Template "Plantilla-Alta-Sec" 1280x800
   Button "Plantilla_6" at 1196,741 size 81x58; TextOff 'Reconocer'; PictureOff "Asleep Check Mark Icon - Sleep Aid Records_2"
      on Press: SetBit("ReconocerTODAS")
      on Release: ResetBit("ReconocerTODAS")
      Appearance <- "AlarmaNueva"
   GraphicView "Plantilla_Visor de gráficos_17" at 4,4 size 87x38; Picture "logo4"
   Button "Plantilla_7" at 479,748 size 78x50; TextOff 'Compres.'
      on Click: ActivateScreen("MTA-CompBAJA", 0)
   Button "Plantilla_8" at 161,748 size 78x50; TextOff 'Torres'
      on Release: ActivateScreen("MTA-TorresCH", 0)
   Button "Plantilla_9" at 81,748 size 78x50; TextOff 'General'; TextOn 'NavigateHome'; PictureOff "NavigateHome_HMI_1"; PictureOn "NavigateHome_HMI_1"
      on Press: ResetBit("VerCh1MTA"); ResetBit("VerCh2MTA"); ResetBit("VerCh3MTA"); ResetBit("VerCh4MTA")
      on Release: ActivateScreen("MTA-Chillers-General", 0)
   Button "Plantilla_12" at 638,748 size 78x50; TextOff 'Luz'; PictureOff "Lamp2_1"
      on Click: ActivateScreen("IluminaciónMTA", 0)
      Appearance <- "MantenerON"
   Button "Plantilla_13" at 400,748 size 78x50; TextOff 'Torres'
      on Click: ActivateScreen("MTA-TorresCAV", 0)
   Button "Plantilla_14" at 321,748 size 78x50; TextOff 'Secadores'
      on Click: ActivateScreen("MTA-SecALTA", 0)
   Button "Plantilla_15" at 558,748 size 78x50; TextOff 'Secadores'
      on Click: ActivateScreen("MTA-SecBaja", 0)
   Button "Plantilla_16" at 241,748 size 78x50; TextOff 'Compres.'
      on Click: ActivateScreen("MTA-CompALTA", 0)
   Button "Plantilla_17" at 1,740 size 78x58; TextOff 'NavigateHome'; PictureOff "NavigateHome_HMI_1"; PictureOn "NavigateHome_HMI_1"
      on Release: ActivateScreen("INICIO", 0)
   GraphicView "Plantilla_Visor de gráficos_1" at 80,740 size 78x6; Picture "indGris"
   GraphicView "Plantilla_Visor de gráficos_2" at 160,740 size 78x6; Picture "indGris"
   GraphicView "Plantilla_Visor de gráficos_3" at 478,740 size 78x6; Picture "indGris"
   GraphicView "Plantilla_Visor de gráficos_4" at 240,740 size 78x6; Picture "indGris"
   GraphicView "Plantilla_Visor de gráficos_5" at 557,740 size 78x6; Picture "indGris"
   GraphicView "Plantilla_Visor de gráficos_6" at 320,740 size 78x6; Picture "indGris"
   GraphicView "Plantilla_Visor de gráficos_7" at 399,740 size 78x6; Picture "indGris"
   GraphicView "Plantilla_Visor de gráficos_11" at 637,740 size 78x6; Picture "indGris"
   GraphicView "Plantilla_Visor de gráficos_8" at 80,740 size 78x6; Picture "indAmarillo"
      Visibility <- "IndCh"
   GraphicView "Plantilla_Visor de gráficos_9" at 160,740 size 78x6; Picture "indAmarillo"
      Visibility <- "IndTrCh"
   GraphicView "Plantilla_Visor de gráficos_10" at 478,740 size 78x6; Picture "indAmarillo"
      Visibility <- "IndCmpBaja"
   GraphicView "Plantilla_Visor de gráficos_12" at 240,740 size 78x6; Picture "indAmarillo"
      Visibility <- "IndCmpAlta"
   GraphicView "Plantilla_Visor de gráficos_13" at 557,740 size 78x6; Picture "indAmarillo"
      Visibility <- "IndSecBaja"
   GraphicView "Plantilla_Visor de gráficos_14" at 320,740 size 78x6; Picture "indAmarillo"
      Visibility <- "IndSecAlta"
   GraphicView "Plantilla_Visor de gráficos_15" at 399,740 size 78x6; Picture "indAmarillo"
      Visibility <- "IndTrCav"
   GraphicView "Plantilla_Visor de gráficos_16" at 637,740 size 78x6; Picture "indAmarillo"
      Visibility <- "MantenerON"
   TextField "Plantilla_Campo de texto_2" at 521,711 size 69x18; Text 'Baja Presión'
   TextField "Plantilla_Campo de texto_4" at 323,711 size 68x18; Text 'Alta Presión'
   TextField "Plantilla_Campo de texto_3" at 139,711 size 40x18; Text 'Chillers'
   Button "Plantilla_3" at 717,748 size 78x50; TextOff 'Text'; PictureOff "Rayo"
      on Click: ActivateScreen("SentronPAC-MTA", 0)
   Button "Plantilla_5" at 957,748 size 78x50; TextOff 'Text'
   Button "Plantilla_11" at 797,748 size 78x50; TextOff 'Variables Analóg.'
      on Click: ActivateScreen("Grafica", 0)
   GraphicView "Plantilla_Visor de gráficos_18" at 717,740 size 78x6; Picture "indGris"
   GraphicView "Plantilla_Visor de gráficos_19" at 797,740 size 78x6; Picture "indGris"
   GraphicView "Plantilla_Visor de gráficos_20" at 877,740 size 78x6; Picture "indGris"
   GraphicView "Plantilla_Visor de gráficos_21" at 957,740 size 78x6; Picture "indGris"
   GraphicView "Plantilla_Visor de gráficos_22" at 1037,740 size 78x6; Picture "indGris"
   GraphicView "Plantilla_Visor de gráficos_23" at 1037,740 size 78x6; Picture "indAmarillo"
      Visibility <- "AnularSirenaCav"
   Button "Plantilla_1" at 1037,749 size 78x50; TextOff 'Anular Sirena'
      on Click: SetBit("AnularSirena?")
   Button "Plantilla_2" at 1117,741 size 78x58; TextOff 'Avisos'
      on Click: ActivateScreen("MTA-Avisos", 0)
   Button "Plantilla_4" at 877,748 size 78x50; TextOff 'Text'
   GraphicView "Plantilla_Visor de gráficos_24" at 877,740 size 78x6; Picture "indGris"
   GraphicView "Plantilla_Visor de gráficos_25" at 877,740 size 78x6; Picture "indGris"
      Visibility <- "AlarmaBoosters"
   Group "Group" at 1,716 size 1276x84
   GraphicView "Plantilla_Visor de gráficos_26" at 68,9 size 91x26; Picture "eProC logo 4 b"
   GraphicView "Plantilla_Visor de gráficos_27" at 9,8 size 49x29; Picture "eProC logo 4 a"
   GraphicIOField "Campo ES gráfico_4" at 981,258 size 280x222; PictureList "Secador1"
      ProcessValue <- "AnimaMS050"
   GraphicView "Visor de gráficos_4" at 999,137 size 234x314; Picture "secador4"
   GraphicView "Visor de gráficos_15" at 999,137 size 234x314; Picture "secador4d_1"
      Visibility <- "MantMS050"
   GraphicIOField "Campo ES gráfico_8" at 571,212 size 366x99; PictureList "Secador2"
      ProcessValue <- "AnimaMS053"
   GraphicView "Visor de gráficos_3" at 592,100 size 363x184; Picture "secador2_3"
   GraphicView "Visor de gráficos_5" at 592,100 size 363x184; Picture "secador2m_1"
      Visibility <- "MantMS053"
   GraphicIOField "Campo ES gráfico_7" at 674,357 size 309x81; PictureList "Secador2"
      ProcessValue <- "AnimaMS052"
   GraphicView "Visor de gráficos_2" at 696,255 size 292x158; Picture "secador3_1"
   GraphicView "Visor de gráficos_6" at 695,255 size 294x158; Picture "secador3d_1"
      Visibility <- "MantMS052"
   GraphicIOField "Campo ES gráfico_6" at 765,490 size 338x86; PictureList "Secador2"
      ProcessValue <- "AnimaMS051"
   GraphicView "Visor de gráficos_1" at 786,405 size 292x142; Picture "secador3_3"
   GraphicView "Visor de gráficos_14" at 786,405 size 292x142; Picture "secador3d_2"
      Visibility <- "MantMS051"
   Rectangle "Plantilla_Rectángulo_1" at 1,716 size 1276x84
      Visibility <- "AnularSirena?"
   TextField "Plantilla_Campo de texto_5" at 32,732 size 696x50; Text '¿Está seguro de ANULAR la sirena? Si decide anular el sistema dejará de emitir avisos sonoros de manera permanente'
      Visibility <- "AnularSirena?"
   Button "Plantilla_Botón_1" at 1232,724 size 37x34; TextOff 'x'
      on Click: ResetBit("AnularSirena?")
      Visibility <- "AnularSirena?"
   Button "Plantilla_Botón_2" at 945,735 size 112x46; TextOff 'Activar'
      on Click: ResetBit("AnularSirenaCav")
      Visibility <- "AnularSirena?"
      Appearance <- "AnularSirenaCav"
   Button "Plantilla_Botón_3" at 1065,735 size 112x46; TextOff 'Desactivar'
      on Click: SetBit("AnularSirenaCav")
      Visibility <- "AnularSirena?"
      Appearance <- "AnularSirenaCav"
   Switch "Interruptor_1" at 640,315 size 40x40; TextOn '1'; TextOff '0'; CaptionText 'Switch'; PictureOff "MECH2"; PictureOn "MECH1"
      ProcessValue <- "MantMS052"
   Switch "Interruptor_2" at 731,440 size 40x40; TextOn '1'; TextOff '0'; CaptionText 'Switch'; PictureOff "MECH2"; PictureOn "MECH1"
      ProcessValue <- "MantMS051"
   Switch "Interruptor_3" at 540,176 size 40x40; TextOn '1'; TextOff '0'; CaptionText 'Switch'; PictureOff "MECH2"; PictureOn "MECH1"
      ProcessValue <- "MantMS053"
   Switch "Interruptor_4" at 1212,488 size 40x40; TextOn '1'; TextOff '0'; CaptionText 'Switch'; PictureOff "MECH2"; PictureOn "MECH1"
      ProcessValue <- "MantMS050"

Template "Plantilla-Baja-Cmp" 1280x800
   Button "Plantilla_6" at 1196,741 size 81x58; TextOff 'Reconocer'; PictureOff "Asleep Check Mark Icon - Sleep Aid Records_2"
      on Press: SetBit("ReconocerTODAS")
      on Release: ResetBit("ReconocerTODAS")
      Appearance <- "AlarmaNueva"
   GraphicView "Plantilla_Visor de gráficos_17" at 4,4 size 87x38; Picture "logo4"
   Button "Plantilla_7" at 479,748 size 78x50; TextOff 'Compres.'
      on Click: ActivateScreen("MTA-CompBAJA", 0)
   Button "Plantilla_8" at 161,748 size 78x50; TextOff 'Torres'
      on Release: ActivateScreen("MTA-TorresCH", 0)
   Button "Plantilla_9" at 81,748 size 78x50; TextOff 'General'; TextOn 'NavigateHome'; PictureOff "NavigateHome_HMI_1"; PictureOn "NavigateHome_HMI_1"
      on Press: ResetBit("VerCh1MTA"); ResetBit("VerCh2MTA"); ResetBit("VerCh3MTA"); ResetBit("VerCh4MTA")
      on Release: ActivateScreen("MTA-Chillers-General", 0)
   Button "Plantilla_12" at 638,748 size 78x50; TextOff 'Luz'; PictureOff "Lamp2_1"
      on Click: ActivateScreen("IluminaciónMTA", 0)
      Appearance <- "MantenerON"
   Button "Plantilla_13" at 400,748 size 78x50; TextOff 'Torres'
      on Click: ActivateScreen("MTA-TorresCAV", 0)
   Button "Plantilla_14" at 321,748 size 78x50; TextOff 'Secadores'
      on Click: ActivateScreen("MTA-SecALTA", 0)
   Button "Plantilla_15" at 558,748 size 78x50; TextOff 'Secadores'
      on Click: ActivateScreen("MTA-SecBaja", 0)
   Button "Plantilla_16" at 241,748 size 78x50; TextOff 'Compres.'
      on Click: ActivateScreen("MTA-CompALTA", 0)
   Button "Plantilla_17" at 1,740 size 78x58; TextOff 'NavigateHome'; PictureOff "NavigateHome_HMI_1"; PictureOn "NavigateHome_HMI_1"
      on Release: ActivateScreen("INICIO", 0)
   GraphicView "Plantilla_Visor de gráficos_1" at 80,740 size 78x6; Picture "indGris"
   GraphicView "Plantilla_Visor de gráficos_2" at 160,740 size 78x6; Picture "indGris"
   GraphicView "Plantilla_Visor de gráficos_3" at 478,740 size 78x6; Picture "indGris"
   GraphicView "Plantilla_Visor de gráficos_4" at 240,740 size 78x6; Picture "indGris"
   GraphicView "Plantilla_Visor de gráficos_5" at 557,740 size 78x6; Picture "indGris"
   GraphicView "Plantilla_Visor de gráficos_6" at 320,740 size 78x6; Picture "indGris"
   GraphicView "Plantilla_Visor de gráficos_7" at 399,740 size 78x6; Picture "indGris"
   GraphicView "Plantilla_Visor de gráficos_11" at 637,740 size 78x6; Picture "indGris"
   GraphicView "Plantilla_Visor de gráficos_8" at 80,740 size 78x6; Picture "indAmarillo"
      Visibility <- "IndCh"
   GraphicView "Plantilla_Visor de gráficos_9" at 160,740 size 78x6; Picture "indAmarillo"
      Visibility <- "IndTrCh"
   GraphicView "Plantilla_Visor de gráficos_10" at 478,740 size 78x6; Picture "indAmarillo"
      Visibility <- "IndCmpBaja"
   GraphicView "Plantilla_Visor de gráficos_12" at 240,740 size 78x6; Picture "indAmarillo"
      Visibility <- "IndCmpAlta"
   GraphicView "Plantilla_Visor de gráficos_13" at 557,740 size 78x6; Picture "indAmarillo"
      Visibility <- "IndSecBaja"
   GraphicView "Plantilla_Visor de gráficos_14" at 320,740 size 78x6; Picture "indAmarillo"
      Visibility <- "IndSecAlta"
   GraphicView "Plantilla_Visor de gráficos_15" at 399,740 size 78x6; Picture "indAmarillo"
      Visibility <- "IndTrCav"
   GraphicView "Plantilla_Visor de gráficos_16" at 637,740 size 78x6; Picture "indAmarillo"
      Visibility <- "MantenerON"
   TextField "Plantilla_Campo de texto_2" at 521,711 size 69x18; Text 'Baja Presión'
   TextField "Plantilla_Campo de texto_4" at 323,711 size 68x18; Text 'Alta Presión'
   TextField "Plantilla_Campo de texto_3" at 139,711 size 40x18; Text 'Chillers'
   Button "Plantilla_3" at 717,748 size 78x50; TextOff 'Text'; PictureOff "Rayo"
      on Click: ActivateScreen("SentronPAC-MTA", 0)
   Button "Plantilla_5" at 957,748 size 78x50; TextOff 'Text'
   Button "Plantilla_11" at 797,748 size 78x50; TextOff 'Variables Analóg.'
      on Click: ActivateScreen("Grafica", 0)
   GraphicView "Plantilla_Visor de gráficos_18" at 717,740 size 78x6; Picture "indGris"
   GraphicView "Plantilla_Visor de gráficos_19" at 797,740 size 78x6; Picture "indGris"
   GraphicView "Plantilla_Visor de gráficos_20" at 877,740 size 78x6; Picture "indGris"
   GraphicView "Plantilla_Visor de gráficos_21" at 957,740 size 78x6; Picture "indGris"
   GraphicView "Plantilla_Visor de gráficos_22" at 1037,740 size 78x6; Picture "indGris"
   GraphicView "Plantilla_Visor de gráficos_23" at 1037,740 size 78x6; Picture "indAmarillo"
      Visibility <- "AnularSirenaCav"
   Button "Plantilla_1" at 1037,749 size 78x50; TextOff 'Anular Sirena'
      on Click: SetBit("AnularSirena?")
   Button "Plantilla_2" at 1117,741 size 78x58; TextOff 'Avisos'
      on Click: ActivateScreen("MTA-Avisos", 0)
   Button "Plantilla_4" at 877,748 size 78x50; TextOff 'Text'
   GraphicView "Plantilla_Visor de gráficos_24" at 877,740 size 78x6; Picture "indGris"
   GraphicView "Plantilla_Visor de gráficos_25" at 877,740 size 78x6; Picture "indGris"
      Visibility <- "AlarmaBoosters"
   Group "Group" at 1,716 size 1276x84
   GraphicView "Plantilla_Visor de gráficos_26" at 68,9 size 91x26; Picture "eProC logo 4 b"
   GraphicView "Plantilla_Visor de gráficos_27" at 9,8 size 49x29; Picture "eProC logo 4 a"
   GraphicIOField "Campo ES gráfico_10" at 491,153 size 189x58; PictureList "BaseSullChico"
      ProcessValue <- "AnimaMC064"
   GraphicIOField "Campo ES gráfico_9" at 427,241 size 189x58; PictureList "BaseSullChico"
      ProcessValue <- "AnimaMC063"
   GraphicIOField "Campo ES gráfico_7" at 387,316 size 178x52; PictureList "BaseSullChico"
      ProcessValue <- "AnimaMC062"
   GraphicIOField "Campo ES gráfico_6" at 340,387 size 178x52; PictureList "BaseSullChico"
      ProcessValue <- "AnimaMC061"
   GraphicIOField "Campo ES gráfico_8" at 275,454 size 197x58; PictureList "BaseSullChico"
      ProcessValue <- "AnimaMC060"
   GraphicView "Visor de gráficos_1" at 467,72 size 269x127; Picture "Baja1X_1"
   GraphicView "Visor de gráficos_7" at 467,72 size 269x127; Picture "Baja1Xd"
      Visibility <- "MantM064"
   GraphicView "Visor de gráficos_2" at 403,160 size 269x127; Picture "Baja1X_1"
   GraphicView "Visor de gráficos_8" at 403,160 size 269x127; Picture "Baja1Xd"
      Visibility <- "MantM063"
   GraphicView "Visor de gráficos_3" at 315,232 size 269x127; Picture "baja2X_2"
   GraphicView "Visor de gráficos_9" at 315,232 size 269x127; Picture "baja2Xd_1"
      Visibility <- "MantM062"
   GraphicView "Visor de gráficos_4" at 267,304 size 269x127; Picture "baja2X_2"
   GraphicView "Visor de gráficos_10" at 267,304 size 269x127; Picture "baja2Xd_1"
      Visibility <- "MantM061"
   GraphicView "Visor de gráficos_5" at 243,376 size 213x127; Picture "baja3X_2"
   GraphicView "Visor de gráficos_11" at 243,376 size 213x127; Picture "baja3Xd"
      Visibility <- "MantM060"
   GraphicView "Visor de gráficos_6" at 132,415 size 202x177; Picture "tanque2X_2"
   IOField "Campo ES_1" at 161,449 size 148x28; FormatPattern s999.9; Unit  bar
      ProcessValue <- "PresiónBAJA"
   GraphicView "Visor de gráficos_12" at 18,528 size 229x141; Picture "Booster-A"
   GraphicIOField "Campo ES gráfico_11" at 68,583 size 48x46; PictureList "Motor Grande"
      ProcessValue <- "AnimaMotBooster"
   GraphicIOField "Campo ES gráfico_12" at 160,500 size 17x32; PictureList "Motor Chico"
      ProcessValue <- "AnimaMotBooster"
   GraphicIOField "Campo ES gráfico_13" at 40,563 size 169x87; PictureList "Hélice"
      ProcessValue <- "Booster_Conf_Marcha"
   GraphicView "Visor de gráficos_18" at 440,520 size 40x40; Picture "MECH2"
   GraphicView "Visor de gráficos_19" at 440,520 size 40x40; Picture "MECH1"
      Visibility <- "Booster2_ModoManten"
   Button "Botón_11" at 440,520 size 40x40; TextOff 'Text'; PictureList "Mantenimiento"
      on Release: SetBit("Booster2_PlsManten")
   GraphicView "Visor de gráficos_17" at 226,528 size 229x141; Picture "Booster-A"
   GraphicIOField "Campo ES gráfico_15" at 286,586 size 48x47; PictureList "Motor Grande"
      ProcessValue <- "AnimaMotBooster2"
   GraphicIOField "Campo ES gráfico_16" at 368,500 size 18x34; PictureList "Motor Chico"
      ProcessValue <- "AnimaMotBooster2"
   GraphicIOField "Campo ES gráfico_17" at 261,565 size 156x84; PictureList "Hélice"
      ProcessValue <- "Booster2_Conf_Marcha"
   GraphicView "Visor de gráficos_13" at 37,520 size 40x40; Picture "MECH2"
   GraphicView "Visor de gráficos_14" at 37,520 size 40x40; Picture "MECH1"
      Visibility <- "Booster_ModoManten"
   Button "Botón_6" at 37,520 size 40x40; TextOff 'Text'; PictureList "Mantenimiento"
      on Release: SetBit("Booster_PlsManten")
   TextField "Campo de texto_4" at 48,674 size 122x19; Text 'Prioridad Marcha'
      Visibility <- "PrioridadBoost1"
   TextField "Campo de texto_10" at 251,674 size 122x19; Text 'Prioridad Marcha'
      Visibility <- "PrioridadBoost2"
   Rectangle "Plantilla_Rectángulo_1" at 1,716 size 1276x84
      Visibility <- "AnularSirena?"
   TextField "Plantilla_Campo de texto_5" at 32,732 size 696x50; Text '¿Está seguro de ANULAR la sirena? Si decide anular el sistema dejará de emitir avisos sonoros de manera permanente'
      Visibility <- "AnularSirena?"
   Button "Plantilla_Botón_1" at 1232,724 size 37x34; TextOff 'x'
      on Click: ResetBit("AnularSirena?")
      Visibility <- "AnularSirena?"
   Button "Plantilla_Botón_2" at 945,735 size 112x46; TextOff 'Activar'
      on Click: ResetBit("AnularSirenaCav")
      Visibility <- "AnularSirena?"
      Appearance <- "AnularSirenaCav"
   Button "Plantilla_Botón_3" at 1065,735 size 112x46; TextOff 'Desactivar'
      on Click: SetBit("AnularSirenaCav")
      Visibility <- "AnularSirena?"
      Appearance <- "AnularSirenaCav"
   Switch "Interruptor_6" at 313,243 size 40x40; TextOn '1'; TextOff '0'; CaptionText 'Switch'; PictureOff "MECH2"; PictureOn "MECH1"
      ProcessValue <- "MantM062"
   Switch "Interruptor_7" at 265,323 size 40x40; TextOn '1'; TextOff '0'; CaptionText 'Switch'; PictureOff "MECH2"; PictureOn "MECH1"
      ProcessValue <- "MantM061"
   Switch "Interruptor_9" at 365,171 size 40x40; TextOn '1'; TextOff '0'; CaptionText 'Switch'; PictureOff "MECH2"; PictureOn "MECH1"
      ProcessValue <- "MantM063"
   Switch "Interruptor_10" at 429,83 size 40x40; TextOn '1'; TextOff '0'; CaptionText 'Switch'; PictureOff "MECH2"; PictureOn "MECH1"
      ProcessValue <- "MantM064"

Template "Plantilla-Baja-Sec" 1280x800
   Button "Plantilla_6" at 1196,741 size 81x58; TextOff 'Reconocer'; PictureOff "Asleep Check Mark Icon - Sleep Aid Records_2"
      on Press: SetBit("ReconocerTODAS")
      on Release: ResetBit("ReconocerTODAS")
      Appearance <- "AlarmaNueva"
   GraphicView "Plantilla_Visor de gráficos_17" at 4,4 size 87x38; Picture "logo4"
   Button "Plantilla_7" at 479,748 size 78x50; TextOff 'Compres.'
      on Click: ActivateScreen("MTA-CompBAJA", 0)
   Button "Plantilla_8" at 161,748 size 78x50; TextOff 'Torres'
      on Release: ActivateScreen("MTA-TorresCH", 0)
   Button "Plantilla_9" at 81,748 size 78x50; TextOff 'General'; TextOn 'NavigateHome'; PictureOff "NavigateHome_HMI_1"; PictureOn "NavigateHome_HMI_1"
      on Press: ResetBit("VerCh1MTA"); ResetBit("VerCh2MTA"); ResetBit("VerCh3MTA"); ResetBit("VerCh4MTA")
      on Release: ActivateScreen("MTA-Chillers-General", 0)
   Button "Plantilla_12" at 638,748 size 78x50; TextOff 'Luz'; PictureOff "Lamp2_1"
      on Click: ActivateScreen("IluminaciónMTA", 0)
      Appearance <- "MantenerON"
   Button "Plantilla_13" at 400,748 size 78x50; TextOff 'Torres'
      on Click: ActivateScreen("MTA-TorresCAV", 0)
   Button "Plantilla_14" at 321,748 size 78x50; TextOff 'Secadores'
      on Click: ActivateScreen("MTA-SecALTA", 0)
   Button "Plantilla_15" at 558,748 size 78x50; TextOff 'Secadores'
      on Click: ActivateScreen("MTA-SecBaja", 0)
   Button "Plantilla_16" at 241,748 size 78x50; TextOff 'Compres.'
      on Click: ActivateScreen("MTA-CompALTA", 0)
   Button "Plantilla_17" at 1,740 size 78x58; TextOff 'NavigateHome'; PictureOff "NavigateHome_HMI_1"; PictureOn "NavigateHome_HMI_1"
      on Release: ActivateScreen("INICIO", 0)
   GraphicView "Plantilla_Visor de gráficos_1" at 80,740 size 78x6; Picture "indGris"
   GraphicView "Plantilla_Visor de gráficos_2" at 160,740 size 78x6; Picture "indGris"
   GraphicView "Plantilla_Visor de gráficos_3" at 478,740 size 78x6; Picture "indGris"
   GraphicView "Plantilla_Visor de gráficos_4" at 240,740 size 78x6; Picture "indGris"
   GraphicView "Plantilla_Visor de gráficos_5" at 557,740 size 78x6; Picture "indGris"
   GraphicView "Plantilla_Visor de gráficos_6" at 320,740 size 78x6; Picture "indGris"
   GraphicView "Plantilla_Visor de gráficos_7" at 399,740 size 78x6; Picture "indGris"
   GraphicView "Plantilla_Visor de gráficos_11" at 637,740 size 78x6; Picture "indGris"
   GraphicView "Plantilla_Visor de gráficos_8" at 80,740 size 78x6; Picture "indAmarillo"
      Visibility <- "IndCh"
   GraphicView "Plantilla_Visor de gráficos_9" at 160,740 size 78x6; Picture "indAmarillo"
      Visibility <- "IndTrCh"
   GraphicView "Plantilla_Visor de gráficos_10" at 478,740 size 78x6; Picture "indAmarillo"
      Visibility <- "IndCmpBaja"
   GraphicView "Plantilla_Visor de gráficos_12" at 240,740 size 78x6; Picture "indAmarillo"
      Visibility <- "IndCmpAlta"
   GraphicView "Plantilla_Visor de gráficos_13" at 557,740 size 78x6; Picture "indAmarillo"
      Visibility <- "IndSecBaja"
   GraphicView "Plantilla_Visor de gráficos_14" at 320,740 size 78x6; Picture "indAmarillo"
      Visibility <- "IndSecAlta"
   GraphicView "Plantilla_Visor de gráficos_15" at 399,740 size 78x6; Picture "indAmarillo"
      Visibility <- "IndTrCav"
   GraphicView "Plantilla_Visor de gráficos_16" at 637,740 size 78x6; Picture "indAmarillo"
      Visibility <- "MantenerON"
   TextField "Plantilla_Campo de texto_2" at 521,711 size 69x18; Text 'Baja Presión'
   TextField "Plantilla_Campo de texto_4" at 323,711 size 68x18; Text 'Alta Presión'
   TextField "Plantilla_Campo de texto_3" at 139,711 size 40x18; Text 'Chillers'
   Button "Plantilla_3" at 717,748 size 78x50; TextOff 'Text'; PictureOff "Rayo"
      on Click: ActivateScreen("SentronPAC-MTA", 0)
   Button "Plantilla_5" at 957,748 size 78x50; TextOff 'Text'
   Button "Plantilla_11" at 797,748 size 78x50; TextOff 'Variables Analóg.'
      on Click: ActivateScreen("Grafica", 0)
   GraphicView "Plantilla_Visor de gráficos_18" at 717,740 size 78x6; Picture "indGris"
   GraphicView "Plantilla_Visor de gráficos_19" at 797,740 size 78x6; Picture "indGris"
   GraphicView "Plantilla_Visor de gráficos_20" at 877,740 size 78x6; Picture "indGris"
   GraphicView "Plantilla_Visor de gráficos_21" at 957,740 size 78x6; Picture "indGris"
   GraphicView "Plantilla_Visor de gráficos_22" at 1037,740 size 78x6; Picture "indGris"
   GraphicView "Plantilla_Visor de gráficos_23" at 1037,740 size 78x6; Picture "indAmarillo"
      Visibility <- "AnularSirenaCav"
   Button "Plantilla_1" at 1037,749 size 78x50; TextOff 'Anular Sirena'
      on Click: SetBit("AnularSirena?")
   Button "Plantilla_2" at 1117,741 size 78x58; TextOff 'Avisos'
      on Click: ActivateScreen("MTA-Avisos", 0)
   Button "Plantilla_4" at 877,748 size 78x50; TextOff 'Text'
   GraphicView "Plantilla_Visor de gráficos_24" at 877,740 size 78x6; Picture "indGris"
   GraphicView "Plantilla_Visor de gráficos_25" at 877,740 size 78x6; Picture "indGris"
   Group "Group" at 1,716 size 1276x84
   GraphicView "Plantilla_Visor de gráficos_26" at 68,9 size 91x26; Picture "eProC logo 4 b"
   GraphicView "Plantilla_Visor de gráficos_27" at 9,8 size 49x29; Picture "eProC logo 4 a"
   GraphicIOField "Campo ES gráfico_1" at 289,314 size 285x90; PictureList "BaseSullChico"
      ProcessValue <- "AnimaMS055"
   GraphicView "Visor de gráficos_2" at 333,200 size 201x179; Picture "secador_1"
   GraphicIOField "Campo ES gráfico_8" at 159,455 size 269x90; PictureList "BaseSullChico"
      ProcessValue <- "AnimaMS054"
   GraphicView "Visor de gráficos_4" at 333,200 size 201x179; Picture "Copia de secador"
      Visibility <- "MantMS055"
   GraphicView "Visor de gráficos_1" at 192,341 size 201x179; Picture "secador_1"
   GraphicView "Visor de gráficos_3" at 192,341 size 201x179; Picture "Copia de secador"
      Visibility <- "MantMS054"
   Rectangle "Plantilla_Rectángulo_1" at 1,716 size 1276x84
      Visibility <- "AnularSirena?"
   TextField "Plantilla_Campo de texto_5" at 32,732 size 696x50; Text '¿Está seguro de ANULAR la sirena? Si decide anular el sistema dejará de emitir avisos sonoros de manera permanente'
      Visibility <- "AnularSirena?"
   Button "Plantilla_Botón_1" at 1232,724 size 37x34; TextOff 'x'
      on Click: ResetBit("AnularSirena?")
      Visibility <- "AnularSirena?"
   Button "Plantilla_Botón_2" at 945,735 size 112x46; TextOff 'Activar'
      on Click: ResetBit("AnularSirenaCav")
      Visibility <- "AnularSirena?"
      Appearance <- "AnularSirenaCav"
   Button "Plantilla_Botón_3" at 1065,735 size 112x46; TextOff 'Desactivar'
      on Click: SetBit("AnularSirenaCav")
      Visibility <- "AnularSirena?"
      Appearance <- "AnularSirenaCav"
   Switch "Interruptor_7" at 271,262 size 40x40; TextOn '1'; TextOff '0'; CaptionText 'Switch'; PictureOff "MECH2"; Authorization "Operación"; PictureOn "MECH1"
      ProcessValue <- "MantMS055"
   Switch "Interruptor_8" at 131,406 size 40x40; TextOn '1'; TextOff '0'; CaptionText 'Switch'; PictureOff "MECH2"; Authorization "Operación"; PictureOn "MECH1"
      ProcessValue <- "MantMS054"

screen "Graf-cau-pot-actual" 1280x800, template "Plantilla"
   TrendView "Visor de curvas_1" at 3,109 size 1268x600
   TextField "Campo de texto_16" at 477,10 size 365x27; Text 'Gráficas - Caudal y Potencia en tiempo real'
   TextField "Campo de texto_1" at 1143,73 size 122x25; Text 'Potencia Kw'
   TextField "Campo de texto_2" at 45,70 size 137x25; Text 'Caudal m3/hs'
   Button "Botón_1" at 271,54 size 150x40; TextOff 'Escalar'
      on Click: ActivateScreen("EcalarSeñAnal", 0)
   Button "Botón_2" at 479,54 size 150x40; TextOff 'Iniciar registro'
      on Click: function_fd9437ed(0, "HistoricoCaudal"); function_fd9437ed(0, "HistoricoPotencia"); SetBit("EstadoRegistro"); function_bb0abc73()
      Appearance <- "EstadoRegistro"
   Button "Botón_3" at 687,54 size 150x40; TextOff 'Parar registro'
      on Click: function_b6526003(0, "HistoricoCaudal"); function_b6526003(0, "HistoricoPotencia"); ResetBit("EstadoRegistro")
   Button "Botón_4" at 895,54 size 150x40; TextOff 'Borrar registro'
      on Click: function_ff1151d2(0, "HistoricoCaudal"); function_ff1151d2(0, "HistoricoPotencia"); ResetBit("EstadoRegistro")

screen "EcalarSeñAnal" 1280x800, template "Plantilla"
   TextField "Campo de texto_1" at 69,133 size 223x27; Text 'Escalar lectura de Caudal:'
   TextField "Campo de texto_2" at 69,375 size 236x27; Text 'Escalar lectura de Potencia:'
   IOField "Campo ES_1" at 415,204 size 119x32; FormatPattern 99999.9
      ProcessValue <- "HI_caudal"
   IOField "Campo ES_2" at 415,274 size 119x32; FormatPattern 99999.9
      ProcessValue <- "LO_caudal"
   IOField "Campo ES_4" at 415,451 size 119x32; FormatPattern 99999.9
      ProcessValue <- "HI_potencia"
   IOField "Campo ES_3" at 415,522 size 119x32; FormatPattern 99999.9
      ProcessValue <- "LO_potencia"
   TextField "Campo de texto_3" at 234,204 size 127x27; Text 'Limite superior'
   TextField "Campo de texto_4" at 234,274 size 118x27; Text 'Limite inferior'
   TextField "Campo de texto_5" at 234,451 size 127x27; Text 'Limite superior'
   TextField "Campo de texto_6" at 234,522 size 118x27; Text 'Limite inferior'
   Button "Botón_3" at 788,329 size 240x49; TextOff 'Grafico Caudal/Potencia'
      on Click: ActivateScreen("Graf-cau-pot-actual", 0)

screen "Graf-cau-pot-historico" 1280x800, template "Plantilla"
   TrendView "Visor de curvas_1" at 3,109 size 1268x600
   TextField "Campo de texto_16" at 477,10 size 334x27; Text 'Gráficas - Hitórico de Caudal y Potencia'
   TextField "Campo de texto_2" at 29,70 size 137x25; Text 'Caudal m3/hs'
   TextField "Campo de texto_1" at 1143,73 size 122x25; Text 'Potencia Kw'
   TextField "Campo de texto_3" at 1143,73 size 122x25; Text 'Potencia Kw'
*)